// TIA Portal project "Industry 4.0_Plant_Logic" (V16) (continued)
REGION Network 1: Filling Process from Tank1
   // When bottle is detected at filling Station, after 2 sec, Tank 01 outlet valve is opened and Pump motor is started.
   // 
   // Tank 01 Outlet valve is closed when defined Liquid A percentage is filled in the bottle.
   // 
   // Liquid A filled value is then moved into Database for Storing purpose.
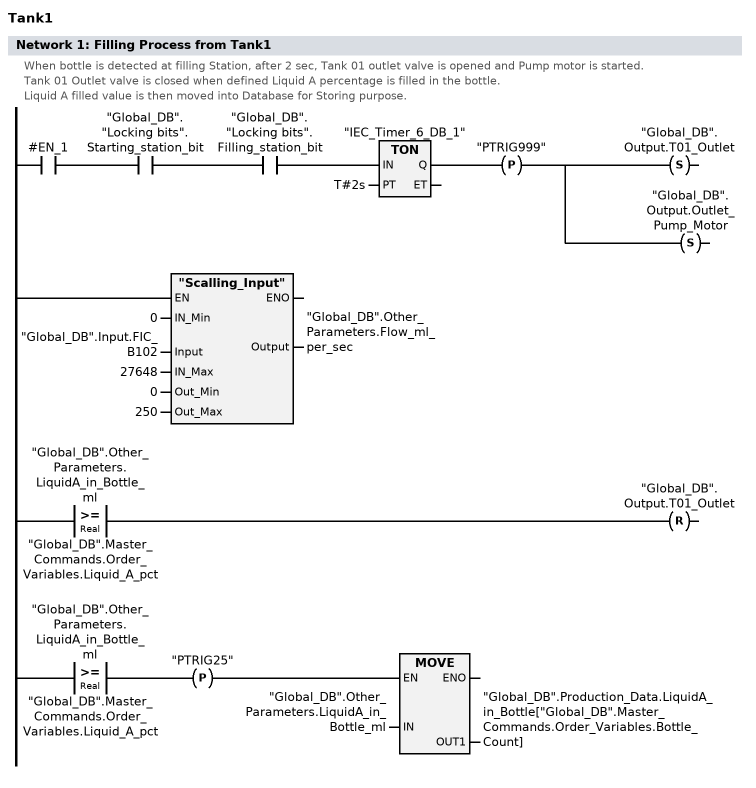
   "IEC_Timer_6_DB_1".TON(IN := #EN_1 AND "Global_DB"."Locking bits".Starting_station_bit AND "Global_DB"."Locking bits".Filling_station_bit,
                          PT := T#2s);
   #_w1 := "IEC_Timer_6_DB_1".Q AND NOT "PTRIG999";   // rising edge
   "PTRIG999" := "IEC_Timer_6_DB_1".Q;
   IF #_w1 THEN
       "Global_DB".Output.T01_Outlet := TRUE;
       "Global_DB".Output.Outlet_Pump_Motor := TRUE;
   END_IF;
   "Scalling_Input"(IN_Min := 0,
                    Input := "Global_DB".Input.FIC_B102,
                    IN_Max := 27648,
                    Out_Min := 0,
                    Out_Max := 250,
                    Output => "Global_DB".Other_Parameters.Flow_ml_per_sec);
   IF "Global_DB".Other_Parameters.LiquidA_in_Bottle_ml >= "Global_DB".Master_Commands.Order_Variables.Liquid_A_pct THEN
       "Global_DB".Output.T01_Outlet := FALSE;
   END_IF;
   #_w2 := "Global_DB".Other_Parameters.LiquidA_in_Bottle_ml >= "Global_DB".Master_Commands.Order_Variables.Liquid_A_pct;
   #_w3 := #_w2 AND NOT "PTRIG25";   // rising edge
   "PTRIG25" := #_w2;
   IF #_w3 THEN
       "Global_DB".Production_Data.LiquidA_in_Bottle["Global_DB".Master_Commands.Order_Variables.Bottle_Count] := "Global_DB".Other_Parameters.LiquidA_in_Bottle_ml;
   END_IF;
END_REGION
END_FUNCTION_BLOCK

FUNCTION_BLOCK "Tank2"   // FB5, LAD
{ S7_Optimized_Access := 'TRUE' }
VERSION : 0.1
   VAR_INPUT
      EN_2 : Bool;
   END_VAR
   VAR_TEMP   // added for the SCL form of the ladder/FBD networks
      _w1 : Bool;
      _w2 : Bool;
      _w3 : Bool;
   END_VAR
BEGIN

REGION Network 1: Tank02 Outlet Solenoid Valve
   // When bottle is filled with liquid A, after 3 sec, Tank 02 outlet valve is opened and Pump motor is started to fill liquid B.
   // 
   // Tank 02 Outlet valve is closed when defined Liquid B percentage is filled in the bottle.
   // 
   // Liquid B filled value is then moved into Database for Storing purpose.
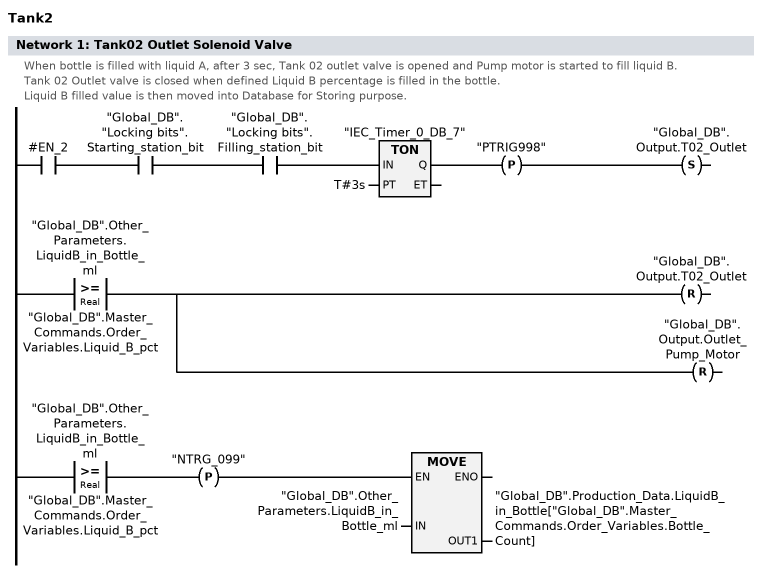
   "IEC_Timer_0_DB_7".TON(IN := #EN_2 AND "Global_DB"."Locking bits".Starting_station_bit AND "Global_DB"."Locking bits".Filling_station_bit,
                          PT := T#3s);
   #_w1 := "IEC_Timer_0_DB_7".Q AND NOT "PTRIG998";   // rising edge
   "PTRIG998" := "IEC_Timer_0_DB_7".Q;
   IF #_w1 THEN "Global_DB".Output.T02_Outlet := TRUE; END_IF;
   IF "Global_DB".Other_Parameters.LiquidB_in_Bottle_ml >= "Global_DB".Master_Commands.Order_Variables.Liquid_B_pct THEN
       "Global_DB".Output.T02_Outlet := FALSE;
       "Global_DB".Output.Outlet_Pump_Motor := FALSE;
   END_IF;
   #_w2 := "Global_DB".Other_Parameters.LiquidB_in_Bottle_ml >= "Global_DB".Master_Commands.Order_Variables.Liquid_B_pct;
   #_w3 := #_w2 AND NOT "NTRG_099";   // rising edge
   "NTRG_099" := #_w2;
   IF #_w3 THEN
       "Global_DB".Production_Data.LiquidB_in_Bottle["Global_DB".Master_Commands.Order_Variables.Bottle_Count] := "Global_DB".Other_Parameters.LiquidB_in_Bottle_ml;
   END_IF;
END_REGION
END_FUNCTION_BLOCK

FUNCTION_BLOCK "ProductionData_Reset"   // FB6, SCL
{ S7_Optimized_Access := 'TRUE' }
VERSION : 0.1
BEGIN

   // when number of filled bottles = Ordered bottle
   // reset the production data buffer and flag order completed To TRUE

   IF "Global_DB".Master_Commands.Order_Variables.Bottle_Count > "Global_DB".Master_Commands.Order_Variables.Quantity THEN
       FOR "Global_DB".Other_Parameters.index := 1 TO 5 BY 1 DO
           "Global_DB".Production_Data.Total_Liquid_in_Bottle["Global_DB".Other_Parameters.index] := 0.0;
           "Global_DB".Production_Data.LiquidA_in_Bottle["Global_DB".Other_Parameters.index] := 0.0;
           "Global_DB".Production_Data.LiquidB_in_Bottle["Global_DB".Other_Parameters.index] := 0.0;
       END_FOR;
       "Global_DB".Master_Commands.Order_Variables.Order_completed := True;
    END_IF;

    // when order is complete, reset the order data

   IF "Global_DB".Master_Commands.Order_Variables.Order_completed = True THEN
       "Global_DB".Master_Commands.Order_Variables.Bottle_Count := 1;
       "Global_DB".Master_Commands.Order_Variables.Order_ID := 0;
       "Global_DB".Master_Commands.Order_Variables.Quantity := 0;
       "Global_DB".Master_Commands.Order_Variables.Liquid_A_pct := 0;
       "Global_DB".Master_Commands.Order_Variables.Liquid_B_pct := 0;
       "Global_DB".Master_Commands.Order_Variables.Order_received := FALSE;
       // "Global_DB".Master_Commands.Order_Variables.Order_completed := FALSE;
   END_IF;
END_FUNCTION_BLOCK

FUNCTION_BLOCK "Reseting_order"   // FB7, SCL
{ S7_Optimized_Access := 'TRUE' }
VERSION : 0.1
BEGIN
   // when next order is received, turn Order_completed flag to FALSE

   "R_TRIG_DB"(CLK := "Global_DB".Master_Commands.Order_Variables.Order_received);

   IF "R_TRIG_DB".Q THEN
       "Global_DB".Master_Commands.Order_Variables.Order_completed := FALSE;
   END_IF;
END_FUNCTION_BLOCK

FUNCTION_BLOCK "Operation_cycle"   // FB8, LAD
{ S7_Optimized_Access := 'TRUE' }
VERSION : 0.1
   VAR
      begun : Bool;
   END_VAR
   VAR_TEMP
      ons1 : Bool;
   END_VAR
   VAR_TEMP   // added for the SCL form of the ladder/FBD networks
      _w1 : Bool;
      _w2 : Bool;
      _w3 : Bool;
   END_VAR
BEGIN

REGION Network 1: Calculate Operation time for one bottle filling and storing in Database for every bottle
   // Operation begin - robot has picked bottle
   // Operation finished - bottle if capped and placed by robot
   // 
   // Note : currently these variables are not getting real-feedback from robots. These are for just simulation.
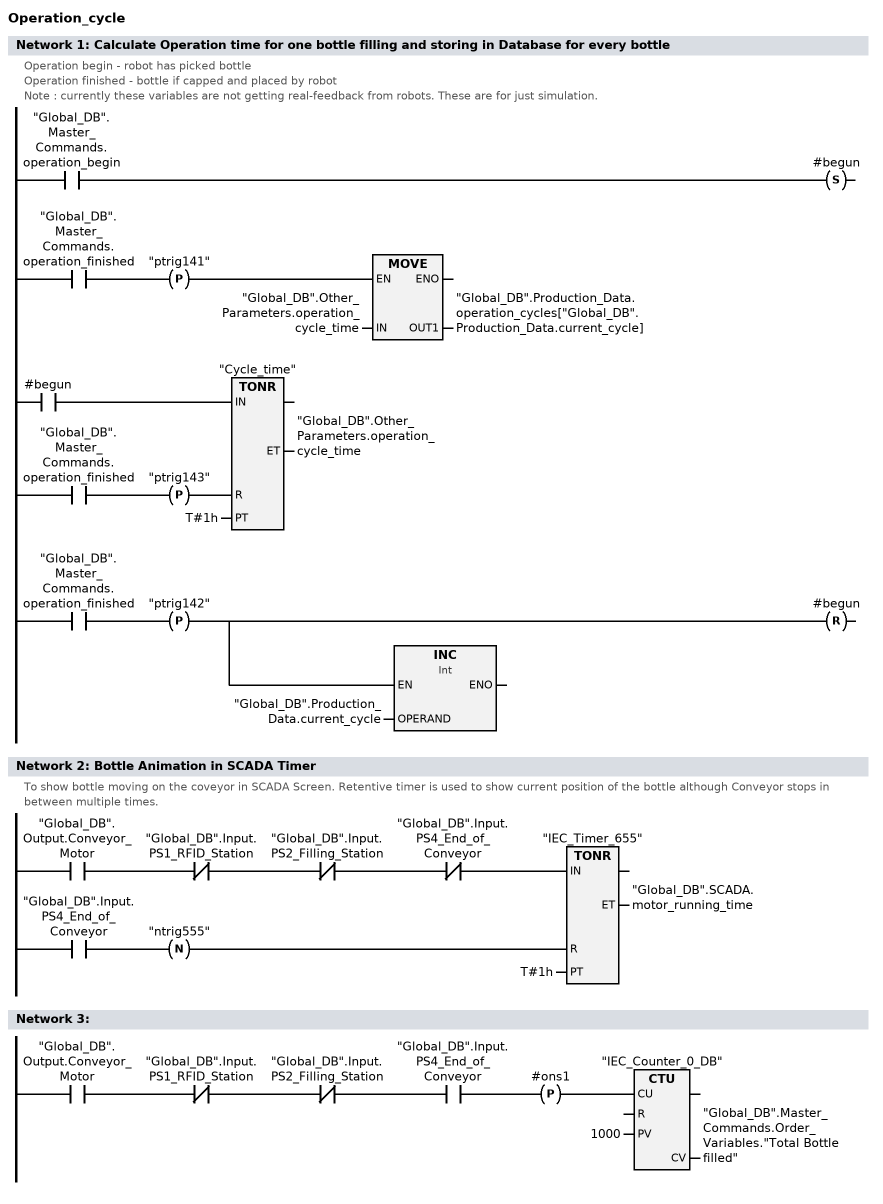
   IF "Global_DB".Master_Commands.operation_begin THEN #begun := TRUE; END_IF;
   #_w1 := "Global_DB".Master_Commands.operation_finished AND NOT "ptrig141";   // rising edge
   "ptrig141" := "Global_DB".Master_Commands.operation_finished;
   IF #_w1 THEN
       "Global_DB".Production_Data.operation_cycles["Global_DB".Production_Data.current_cycle] := "Global_DB".Other_Parameters.operation_cycle_time;
   END_IF;
   #_w2 := "Global_DB".Master_Commands.operation_finished AND NOT "ptrig143";   // rising edge
   "ptrig143" := "Global_DB".Master_Commands.operation_finished;
   "Cycle_time".TONR(IN := #begun,
                     R := #_w2,
                     PT := T#1h,
                     ET => "Global_DB".Other_Parameters.operation_cycle_time);
   #_w3 := "Global_DB".Master_Commands.operation_finished AND NOT "ptrig142";   // rising edge
   "ptrig142" := "Global_DB".Master_Commands.operation_finished;
   IF #_w3 THEN
       #begun := FALSE;
       "Global_DB".Production_Data.current_cycle := "Global_DB".Production_Data.current_cycle + 1;
   END_IF;
END_REGION

REGION Network 2: Bottle Animation in SCADA Timer
   // To show bottle moving on the coveyor in SCADA Screen. Retentive timer is used to show current position of the bottle although Conveyor stops in between multiple times.
   #_w1 := NOT "Global_DB".Input.PS4_End_of_Conveyor AND "ntrig555";   // falling edge
   "ntrig555" := "Global_DB".Input.PS4_End_of_Conveyor;
   "IEC_Timer_655".TONR(IN := "Global_DB".Output.Conveyor_Motor AND NOT "Global_DB".Input.PS1_RFID_Station AND NOT "Global_DB".Input.PS2_Filling_Station AND NOT "Global_DB".Input.PS4_End_of_Conveyor,
                        R := #_w1,
                        PT := T#1h,
                        ET => "Global_DB".SCADA.motor_running_time);
END_REGION

REGION Network 3
   #_w1 := "Global_DB".Output.Conveyor_Motor AND NOT "Global_DB".Input.PS1_RFID_Station AND NOT "Global_DB".Input.PS2_Filling_Station AND "Global_DB".Input.PS4_End_of_Conveyor;
   #_w2 := #_w1 AND NOT #ons1;   // rising edge
   #ons1 := #_w1;
   "IEC_Counter_0_DB".CTU(CU := #_w2,
                          PV := 1000,
                          CV => "Global_DB".Master_Commands.Order_Variables."Total Bottle filled");
END_REGION
END_FUNCTION_BLOCK

FUNCTION_BLOCK "Array_Voltage_Logic"   // FB9, SCL
{ S7_Optimized_Access := 'TRUE' }
VERSION : 0.1
BEGIN




       "Global_DB".Array_Voltage["i"] :="Global_DB".Motor_Output_PCT;
       "i" := "i" + 1;
END_FUNCTION_BLOCK

// folder: Functions

FUNCTION "Scalling_Input" : Void   // FC1, FBD
{ S7_Optimized_Access := 'TRUE' }
VERSION : 0.1
   VAR_INPUT
      IN_Min : Int;
      Input : Int;
      IN_Max : Int;
      Out_Min : Int;
      Out_Max : Int;
   END_VAR
   VAR_OUTPUT
      Output : Real;
   END_VAR
   VAR_TEMP
      Normed : Real;
   END_VAR
BEGIN

REGION Network 1
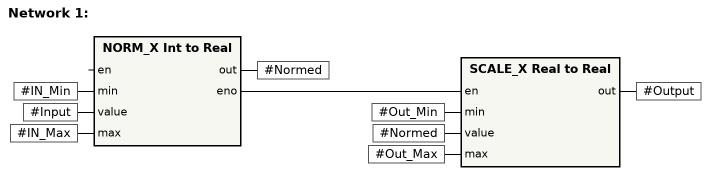
   #Normed := NORM_X(MIN := #IN_Min, VALUE := #Input, MAX := #IN_Max);
   #Output := SCALE_X(MIN := #Out_Min, VALUE := #Normed, MAX := #Out_Max);
END_REGION
END_FUNCTION

FUNCTION "Scalling_Output" : Void   // FC2, FBD
{ S7_Optimized_Access := 'TRUE' }
VERSION : 0.1
   VAR_INPUT
      IN_Min : Int;
      Input : Int;
      IN_Max : Int;
      Out_Min : Int;
      Out_Max : Int;
   END_VAR
   VAR_OUTPUT
      Output : Int;
   END_VAR
   VAR_TEMP
      Normed : Real;
   END_VAR
BEGIN

REGION Network 1
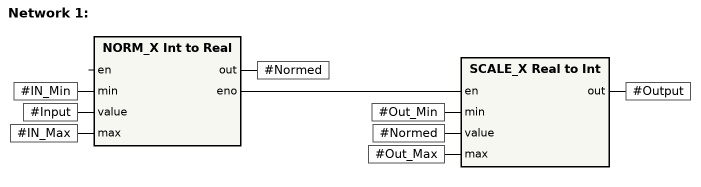
   #Normed := NORM_X(MIN := #IN_Min, VALUE := #Input, MAX := #IN_Max);
   #Output := SCALE_X(MIN := #Out_Min, VALUE := #Normed, MAX := #Out_Max);
END_REGION
END_FUNCTION

FUNCTION "Reading" : Void   // FC3, SCL
{ S7_Optimized_Access := 'TRUE' }
VERSION : 0.1
BEGIN
   // Reading inputs from PLC terminals to Global_DB

   "Global_DB".Input.FIC_B102 := "FIC_B102";
   "Global_DB".Input.LIC_B101 := "LIC_B101";
   "Global_DB".Input.PS1_RFID_Station := "PS1_RFID_Station";
   "Global_DB".Input.PS2_Filling_Station := "PS2_Filling_Station";
   "Global_DB".Input.PS3_Quality_Station := "PS3_Quality_Station";
   "Global_DB".Input.PS4_End_of_Conveyor := "PS4_End_of_Conveyor";
   "Global_DB".Input.T01_Low_Level := "T01_Low_Level";
   "Global_DB".Input.T01_High_Level := "T01_High_Level";
END_FUNCTION

FUNCTION "Writing" : Void   // FC4, SCL
{ S7_Optimized_Access := 'TRUE' }
VERSION : 0.1
BEGIN
   // Writing Output from Global_DB to PLC Terminal

   "T01_Outlet" := "Global_DB".Output.T01_Outlet;
   "T02_Outlet" := "Global_DB".Output.T02_Outlet;

   "Outlet_Pump_Motor" := "Global_DB".Output.Outlet_Pump_Motor;
   "Conveyor_Motor" := "Global_DB".Output.Conveyor_Motor;
END_FUNCTION

FUNCTION "Filling_Logik" : Void   // FC5, LAD
{ S7_Optimized_Access := 'TRUE' }
VERSION : 0.1
   VAR_INPUT
      PS2_Filling_Station : Bool;
      FIC_B102 : Int;
      Liquid_AorB_in_Bottle_ml : Real;
      Liquid_AorB_pct : Int;
      Wait_to_fill : Time;
   END_VAR
   VAR_OUTPUT
      Flow_ml_per_sec : Real;
      FillingData_LiqAorB_ml : Real;
   END_VAR
   VAR_IN_OUT
      Outlet_of_tanks : Bool;
   END_VAR
   VAR_TEMP
      PTRIG1 : Bool;
      PTRIG2 : Bool;
      PTRIG3 : Bool;
      PTRIG4 : Bool;
   END_VAR
BEGIN

REGION Network 1
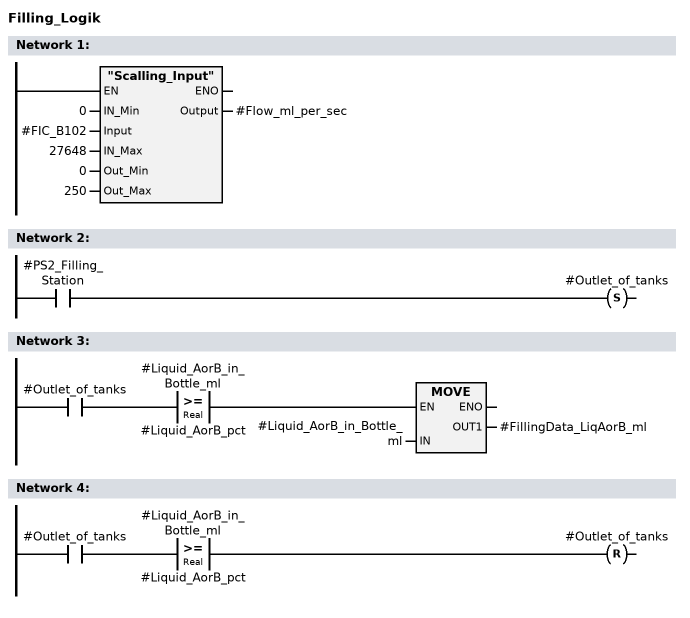
   RUNG wire#powerrail
      "Scalling_Input"(IN_Min := 0, Input := #FIC_B102, IN_Max := 27648, Out_Min := 0, Out_Max := 250, Output => #Flow_ml_per_sec)
   END_RUNG
   // the same network as SCL:
   "Scalling_Input"(IN_Min := 0,
                    Input := #FIC_B102,
                    IN_Max := 27648,
                    Out_Min := 0,
                    Out_Max := 250,
                    Output => #Flow_ml_per_sec);
END_REGION

REGION Network 2
   RUNG wire#powerrail
      Contact( #PS2_Filling_Station )
      S_Coil( #Outlet_of_tanks )
   END_RUNG
   // the same network as SCL:
   IF #PS2_Filling_Station THEN #Outlet_of_tanks := TRUE; END_IF;
END_REGION

REGION Network 3
   RUNG wire#powerrail
      Contact( #Outlet_of_tanks )
      { S7_Templates := "SrcType := Real" } GE_Contact(in1 := #Liquid_AorB_in_Bottle_ml, in2 := #Liquid_AorB_pct)
      Move(in := #Liquid_AorB_in_Bottle_ml, out1 => #FillingData_LiqAorB_ml)
   END_RUNG
   // the same network as SCL:
   IF #Outlet_of_tanks AND (#Liquid_AorB_in_Bottle_ml >= #Liquid_AorB_pct) THEN
       #FillingData_LiqAorB_ml := #Liquid_AorB_in_Bottle_ml;
   END_IF;
END_REGION

REGION Network 4
   RUNG wire#powerrail
      Contact( #Outlet_of_tanks )
      { S7_Templates := "SrcType := Real" } GE_Contact(in1 := #Liquid_AorB_in_Bottle_ml, in2 := #Liquid_AorB_pct)
      R_Coil( #Outlet_of_tanks )
   END_RUNG
   // the same network as SCL:
   IF #Outlet_of_tanks AND (#Liquid_AorB_in_Bottle_ml >= #Liquid_AorB_pct) THEN
       #Outlet_of_tanks := FALSE;
   END_IF;
END_REGION
END_FUNCTION

(* ===== HMI "HMI_RT_1" =====
system functions are stored by id; their names below are inferred from use
connection "PLCs71200": ETHERNET, SMART_S7_1200_OMS
connection "HMI_Connection_1": ETHERNET, SMART_S7_1200_OMS

HMI tags "Default tag table"
   "Conveyor_Motor" : Bool = PLC Global_DB.Output.Conveyor_Motor AT %DB1.DBX6.3, 1 s
   "Outlet_Pump_Motor" : Bool = PLC Global_DB.Output.Outlet_Pump_Motor AT %DB1.DBX6.2, 1 s
   "T01_Outlet_Valve" : Bool = PLC Global_DB.Output.T01_Outlet AT %DB1.DBX6.0, 1 s
   "T02_Outlet_Valve" : Bool = PLC Global_DB.Output.T02_Outlet AT %DB1.DBX6.1, 1 s
   "T02_fluid Low level" : Real = PLC Global_DB.Other_Parameters.T02_Low_Level_Limit AT %DB1.DBD30, 1 s
   "Global_DB_Other_Parameters_Liquid_A_pct" : Int = PLC Global_DB.Master_Commands.Order_Variables.Liquid_A_pct AT %DB1.DBW52, 1 s
   "Global_DB_Other_Parameters_Liquid_B_pct" : Int = PLC Global_DB.Master_Commands.Order_Variables.Liquid_B_pct AT %DB1.DBW54, 1 s
   "Total_Liquid_in_Bottle{0}" : Array [0..4] of Real = PLC Global_DB.Production_Data.Total_Liquid_in_Bottle AT %DB1.DBX66.0, 1 s
   "T02_Low_Level_Limit" : Real = PLC Global_DB.Other_Parameters.T02_Low_Level_Limit AT %DB1.DBD30, 1 s
   "Global_DB_Input_T01_Low_Level" : Bool = PLC Global_DB.Input.T01_Low_Level AT %DB1.DBX4.4, 1 s
   "Global_DB_Input_T01_High_Level" : Bool = PLC Global_DB.Input.T01_High_Level AT %DB1.DBX4.5, 1 s
   "Error_Alarm" : Word = PLC Global_DB.Error.Alarm AT %DB1.DBW42, 1 s
   "Global_DB_Input_FIC_B102" : Int = PLC Global_DB.Input.FIC_B102 AT %DB1.DBW0, 1 s
   "Global_DB_Input_LIC_B101" : Int = PLC Global_DB.Input.LIC_B101 AT %DB1.DBW2, 1 s
   "Global_DB_Production_Data_Bottle_Count" : Int = PLC Global_DB.Master_Commands.Order_Variables.Bottle_Count AT %DB1.DBW58, 1 s
   "Flow_ml_per_sec" : Real = PLC Global_DB.Other_Parameters.Flow_ml_per_sec AT %DB1.DBD10, 1 s
   "PS1_RFID_Station" : Bool = PLC Global_DB.Input.PS1_RFID_Station AT %DB1.DBX4.0, 1 s
   "PS2_Filling_Station" : Bool = PLC Global_DB.Input.PS2_Filling_Station AT %DB1.DBX4.1, 1 s
   "PS3_Quality_Station" : Bool = PLC Global_DB.Input.PS3_Quality_Station AT %DB1.DBX4.2, 1 s
   "PS4_End_of_Conveyor" : Bool = PLC Global_DB.Input.PS4_End_of_Conveyor AT %DB1.DBX4.3, 1 s

discrete alarms
   1: 'Level of Tank01 is high', class Errors, trigger "Global_DB_Error_HIgh level Alarm T01" bit 0
   2: 'Level of Tank01 is low', class Errors, trigger "Global_DB_Error_low level Alarm T01" bit 0

analog alarms
   4: 'Level of Tank02 is high', class Warnings, trigger "Global_DB_Other_Parameters_T02_High_Level_Limit"
   5: 'Level of Tank02 is low', class Warnings, trigger "T02_Low_Level_Limit"

recipe "combinations": Liquid A <- "Global_DB_Other_Parameters_Liquid_A_pct", Liquid B <- "Global_DB_Other_Parameters_Liquid_B_pct"

screen "Different jobs" 800x480
   TextField "Text field_1" at 339,11 size 221x27; Text 'Diffrent Jobs / Gruppe der Ingenieure'
   GraphicView "Graphic view_61" at 2,4 size 149x43; Picture "logo2"
   DateTimeField "Date/time field_1" at 629,14 size 166x19
   Button "Back" at 181,104 size 188x64; TextOn 'Back / Zurück'; TextOff 'Back / Zurück'
      on Release: function_efd93a16()
   Button "Toggle language" at 177,208 size 192x70; TextOn 'Toggle language / Sprache Wechseln'; TextOff 'Toggle language / Sprache Wechseln'
      on Release: function_fb9197e8(-1)
   Button "Online" at 177,320 size 192x66; TextOn 'Online'; TextOff 'Online'
   Button "Offline" at 460,103 size 189x65; TextOn 'Offline'; TextOff 'Offline'
   Button "Stop Runtime" at 460,209 size 189x69; TextOn 'Stop Runtime / Laufzeit anhalten'; TextOff 'Stop Runtime / Laufzeit anhalten'
   Button "Transfer" at 457,320 size 192x65; TextOn 'Transfer / Übertragung'; TextOff 'Transfer / Übertragung'
   Button "Button_1" at 6,432 size 88x38; TextOff 'Root'
      on Release: ActivateScreen("Root screen", 0)
      on Press: ActivateScreen("Root screen", 0)
   Button "Button_2" at 99,432 size 93x38; TextOff 'User / Benutzer'
      on Release: ActivateScreen("User administration", 0)
      on Press: ActivateScreen("User administration", 0)
   Button "Button_3" at 197,431 size 96x39; TextOff 'Alarms / Alarme'
      on Release: ActivateScreen("Alarm screen", 0)
      on Press: ActivateScreen("Alarm screen", 0)
   Button "Button_4" at 298,431 size 121x39; TextOff 'PLC diagnose / SPS Diagnose'
      on Release: ActivateScreen("SIMATIC PLC system diagnostics", 0)
      on Press: ActivateScreen("SIMATIC PLC system diagnostics", 0)
   Button "Button_5" at 425,431 size 106x39; TextOff 'Recipes / Rezepte'
      on Release: ActivateScreen("Recipes management", 0)
      on Press: ActivateScreen("Recipes management", 0)
   Button "Button_6" at 537,431 size 113x39; TextOff 'Visulization / Visulisierung'
      on Release: ActivateScreen("visualization", 0)
      on Press: ActivateScreen("visualization", 0)
   Button "Button_7" at 654,431 size 139x39; TextOff 'Historic Data / Frühere Daten'
      on Release: ActivateScreen("Historical Data", 0)
      on Press: ActivateScreen("Historical Data", 0)

screen "visualization" 800x480
   GraphicView "Graphic view_38" at 637,99 size 155x90; Picture "Graphic_80"
   GraphicView "Graphic view_91" at 719,110 size 19x17; Picture "Graphic_70"
   GraphicView "Graphic view_84" at 735,110 size 19x17; Picture "Graphic_70"
   GraphicView "Graphic view_26" at 751,110 size 19x17; Picture "Graphic_70"
   GraphicView "Graphic view_83" at 768,110 size 19x17; Picture "Graphic_70"
   TextField "Text field_2" at 600,134 size 15x23; Text '4'
   GraphicView "Graphic view_22" at 285,216 size 38x24; Picture "Graphic_43"
   GraphicView "Graphic view_4" at 442,213 size 29x22; Picture "Graphic_60"
   GraphicView "Graphic view_32" at 2,111 size 162x71; Picture "Graphic_76"
   GraphicView "Graphic view_27" at 181,310 size 49x14; Picture "Graphic_65"
   GraphicView "Graphic view_61" at 2,4 size 149x43; Picture "logo2"
   DateTimeField "Date/time field_1" at 629,14 size 167x19
   TextField "Text field_1" at 346,11 size 115x25; Text 'Visulization / Visulisierung'
   Group "Group_1" at 637,99 size 155x90; Picture "Graphic_80"
   GraphicView "Graphic view_72" at 633,201 size 162x71; Picture "Graphic_76"
   GraphicView "Graphic view_82" at 713,205 size 22x17; Picture "Graphic_70"
   GraphicView "Graphic view_85" at 676,205 size 22x17; Picture "Graphic_70"
   GraphicView "Graphic view_87" at 694,205 size 22x17; Picture "Graphic_70"
   GraphicView "Graphic view_93" at 690,211 size 22x17; Picture "Graphic_70"
   GraphicView "Graphic view_103" at 671,211 size 22x17; Picture "Graphic_70"
   Group "Group_4" at 587,131 size 43x28
   GraphicView "Graphic view_89" at 658,205 size 22x17; Picture "Graphic_70"
   GraphicView "Graphic view_86" at 653,211 size 22x17; Picture "Graphic_70"
   GraphicView "Graphic view_92" at 649,217 size 22x17; Picture "Graphic_70"
   GraphicView "Graphic view_90" at 645,222 size 22x17; Picture "Graphic_70"
   GraphicView "Graphic view_80" at 708,211 size 22x17; Picture "Graphic_70"
   GraphicView "Graphic view_1" at 258,95 size 95x94; Picture "Graphic_1"
   GraphicView "Graphic view_21" at 318,221 size 130x14; Picture "Graphic_41"
   GraphicView "Graphic view_2" at 414,97 size 95x94; Picture "Graphic_1"
   GraphicView "Graphic view_11" at 415,100 size 28x90; Picture "Graphic_15"
   GraphicView "Graphic view_12" at 451,187 size 22x16; Picture "Graphic_57"
   GraphicView "Graphic view_19" at 451,201 size 32x16; Picture "Graphic_48"
      Appearance <- "T01_Outlet_Valve"
   GraphicView "Graphic view_5" at 280,61 size 41x122; Picture "Graphic_4"
   GraphicView "Graphic view_9" at 322,236 size 44x38; Picture "Graphic_9"
   GraphicView "Graphic view_7" at 240,214 size 54x28; Picture "Graphic_10"
      Appearance <- "Outlet_Pump_Motor"
   GraphicView "Graphic view_13" at 292,185 size 24x17; Picture "Graphic_57"
   GraphicView "Graphic view_18" at 292,200 size 35x19; Picture "Graphic_48"
      Appearance <- "T02_Outlet_Valve"
   GraphicView "Graphic view_23" at 294,237 size 20x12; Picture "Graphic_57"
   GraphicView "Graphic view_24" at 364,257 size 18x17; Picture "Graphic_63"
   GraphicView "Graphic view_28" at 391,282 size 22x22; Picture "Graphic_72"
   GraphicView "Graphic view_25" at 377,257 size 36x27; Picture "Graphic_64"
   GraphicView "Graphic view_20" at 294,247 size 32x27; Picture "Graphic_62"
   GraphicView "Graphic view_6" at 486,102 size 47x25; Picture "Graphic_5"
      Appearance <- "Global_DB_Input_T01_High_Level"
   GraphicView "Graphic view_8" at 486,170 size 47x25; Picture "Graphic_5"
      Appearance <- "Global_DB_Input_T01_Low_Level"
   IOField "I/O field_1" at 563,220 size 71x32; FormatPattern 999
      ProcessValue <- "Global_DB_Production_Data_Bottle_Count"
   IOField "I/O field_2" at 102,246 size 102x32; FormatPattern 999.99; Unit ml/s
      ProcessValue <- "Flow_ml_per_sec"
   GraphicView "Graphic view_33" at 100,114 size 22x17; Picture "Graphic_70"
   GraphicView "Graphic view_34" at 95,121 size 22x17; Picture "Graphic_70"
   GraphicView "Graphic view_35" at 82,114 size 22x17; Picture "Graphic_70"
   GraphicView "Graphic view_36" at 45,113 size 22x17; Picture "Graphic_70"
   GraphicView "Graphic view_37" at 28,113 size 22x17; Picture "Graphic_70"
   GraphicView "Graphic view_39" at 65,113 size 22x17; Picture "Graphic_70"
   GraphicView "Graphic view_41" at 22,119 size 22x17; Picture "Graphic_70"
   GraphicView "Graphic view_42" at 76,121 size 22x17; Picture "Graphic_70"
   GraphicView "Graphic view_43" at 41,118 size 22x17; Picture "Graphic_70"
   GraphicView "Graphic view_44" at 60,119 size 22x17; Picture "Graphic_70"
   GraphicView "Graphic view_46" at 118,115 size 22x17; Picture "Graphic_70"
   GraphicView "Graphic view_47" at 72,127 size 22x17; Picture "Graphic_70"
   GraphicView "Graphic view_51" at 53,127 size 22x17; Picture "Graphic_70"
   TextField "Text field_4" at 176,132 size 25x23; Text '6 / 14'
   GraphicView "Graphic view_50" at 36,126 size 22x17; Picture "Graphic_70"
   GraphicView "Graphic view_48" at 30,132 size 22x17; Picture "Graphic_70"
   GraphicView "Graphic view_49" at 17,126 size 22x17; Picture "Graphic_70"
   GraphicView "Graphic view_45" at 13,132 size 22x17; Picture "Graphic_70"
   TextField "Text field_3" at 8,250 size 93x23; Text 'Flow Rate:'
   GraphicView "Graphic view_10" at 260,98 size 28x90; Picture "Graphic_15"
   Button "Button_1" at 6,432 size 88x38; TextOff 'Root'
      on Release: ActivateScreen("Root screen", 0)
      on Press: ActivateScreen("Root screen", 0)
   Button "Button_2" at 99,432 size 93x38; TextOff 'User / Benutzer'
      on Release: ActivateScreen("User administration", 0)
      on Press: ActivateScreen("User administration", 0)
   Button "Button_3" at 197,431 size 96x39; TextOff 'Alarms / Alarme'
      on Release: ActivateScreen("Alarm screen", 0)
      on Press: ActivateScreen("Alarm screen", 0)
   Button "Button_4" at 298,431 size 121x39; TextOff 'PLC diagnose / SPS Diagnose'
      on Release: ActivateScreen("SIMATIC PLC system diagnostics", 0)
      on Press: ActivateScreen("SIMATIC PLC system diagnostics", 0)
   Button "Button_5" at 425,431 size 106x39; TextOff 'Recipes / Rezepte'
      on Release: ActivateScreen("Recipes management", 0)
      on Press: ActivateScreen("Recipes management", 0)
   Button "Button_6" at 537,431 size 113x39; TextOff 'Visulization / Visulisierung'
      on Release: ActivateScreen("visualization", 0)
      on Press: ActivateScreen("visualization", 0)
   Button "Button_7" at 654,431 size 139x39; TextOff 'Historic Data / Frühere Daten'
      on Release: ActivateScreen("Historical Data", 0)
      on Press: ActivateScreen("Historical Data", 0)
   GraphicView "Graphic view_68" at 140,388 size 41x27; Picture "Graphic_93"
      Appearance <- "Conveyor_Motor"
   GraphicView "Graphic view_17" at 137,331 size 510x69; Picture "Graphic_28"
   GraphicView "Graphic view_40" at 185,338 size 35x24; Picture "Graphic_88"
   GraphicView "Graphic view_29" at 241,304 size 29x72; Picture "Graphic_70"
      Visibility <- "PS1_RFID_Station"
   GraphicView "Graphic view_15" at 265,306 size 22x41; Picture "Graphic_24"
      Appearance <- "PS1_RFID_Station"
   GraphicView "Graphic view_67" at 323,304 size 29x72; Picture "Graphic_70"
      Visibility <- "PS2_Filling_Station"
   GraphicView "Graphic view_14" at 340,305 size 22x41; Picture "Graphic_24"
      Appearance <- "PS2_Filling_Station"
   GraphicView "Graphic view_3" at 445,307 size 22x41; Picture "Graphic_24"
      Appearance <- "PS3_Quality_Station"
   GraphicView "Graphic view_65" at 423,304 size 29x72; Picture "Graphic_70"
      Visibility <- "PS3_Quality_Station"
   GraphicView "Graphic view_63" at 511,304 size 29x72; Picture "Graphic_70"
      Visibility <- "PS4_End_of_Conveyor"
   GraphicView "Graphic view_16" at 532,307 size 22x41; Picture "Graphic_24"
      Appearance <- "PS4_End_of_Conveyor"

screen "Root screen" 800x480
   TextField "HmiScreenItemData" at 64,85 size 675x54; Text 'Welcome to liquid filling plant based on Industry 4.0 / Willkommen bei der Flüssigkeitsabfüllanlage auf Basis von Industrie 4.0'
   TextField "Text field_1" at 339,10 size 158x27; Text 'Root Screen / Root Bildschirm'
   GraphicView "Graphic view_61" at 2,4 size 149x43; Picture "logo2"
   DateTimeField "Date/time field_1" at 629,14 size 166x19
   Button "Button_8" at 263,167 size 115x69; TextOff 'START'
   Button "Button_9" at 425,166 size 115x69; TextOff 'STOP / STOPP'
   Switch "Switch_1" at 287,262 size 226x63; TextOn 'Emergency is pressed / Notruf wird gedrückt'; CaptionText 'Switch'; TextOff 'Emergency is released / Notfall wird ausgelöst'
   Button "Button_1" at 6,432 size 88x38; TextOff 'Root'
      on Release: ActivateScreen("Root screen", 0)
      on Press: ActivateScreen("Root screen", 0)
   Button "Button_2" at 99,432 size 93x38; TextOff 'User / Benutzer'
      on Release: ActivateScreen("User administration", 0)
      on Press: ActivateScreen("User administration", 0)
   Button "Button_3" at 197,431 size 96x39; TextOff 'Alarms / Alarme'
      on Release: ActivateScreen("Alarm screen", 0)
      on Press: ActivateScreen("Alarm screen", 0)
   Button "Button_4" at 298,431 size 121x39; TextOff 'PLC diagnose / SPS Diagnose'
      on Release: ActivateScreen("SIMATIC PLC system diagnostics", 0)
      on Press: ActivateScreen("SIMATIC PLC system diagnostics", 0)
   Button "Button_5" at 425,431 size 106x39; TextOff 'Recipes / Rezepte'
      on Release: ActivateScreen("Recipes management", 0)
      on Press: ActivateScreen("Recipes management", 0)
   Button "Button_6" at 537,431 size 113x39; TextOff 'Visulization / Visulisierung'
      on Release: ActivateScreen("visualization", 0)
      on Press: ActivateScreen("visualization", 0)
   Button "Button_7" at 654,431 size 139x39; TextOff 'Historic Data / Frühere Daten'
      on Release: ActivateScreen("Historical Data", 0)
      on Press: ActivateScreen("Historical Data", 0)
   Button "Button_12" at 9,156 size 176x46; TextOff 'Different Jobs / System Bildschirme'
      on Release: ActivateScreen("Different jobs", 0)
      on Press: ActivateScreen("Different jobs", 0)
   Button "Button_11" at 16,222 size 157x45; TextOff 'Engineer / Ingenieur'; Authorization "Engineer"
      on Release: ActivateScreen("Engineer Screen", 0)
      on Press: ActivateScreen("Engineer Screen", 0)
   Button "Button_13" at 12,287 size 164x49; TextOff 'Change Langauge / Sprache Wechseln'
      on Click: function_fb9197e8(-1)

screen "User administration" 800x480
   TextField "Text field_1" at 319,10 size 198x27; Text 'User Administration / Benutzerverwaltung'
   GraphicView "Graphic view_61" at 2,4 size 149x43; Picture "logo2"
   DateTimeField "Date/time field_1" at 628,14 size 167x19
   UserView "User view_1" at 9,64 size 781x289
   Button "Button_8" at 10,372 size 134x39; TextOff 'Logoff / Abmeldung'
      on Release: function_f23ef4c9()
      on Press: function_f23ef4c9()
   Button "Button_1" at 6,432 size 88x38; TextOff 'Root'
      on Release: ActivateScreen("Root screen", 0)
      on Press: ActivateScreen("Root screen", 0)
   Button "Button_2" at 99,432 size 93x38; TextOff 'User / Benutzer'
      on Release: ActivateScreen("User administration", 0)
      on Press: ActivateScreen("User administration", 0)
   Button "Button_3" at 197,431 size 96x39; TextOff 'Alarms / Alarme'
      on Release: ActivateScreen("Alarm screen", 0)
      on Press: ActivateScreen("Alarm screen", 0)
   Button "Button_4" at 298,431 size 121x39; TextOff 'PLC diagnose / SPS Diagnose'
      on Release: ActivateScreen("SIMATIC PLC system diagnostics", 0)
      on Press: ActivateScreen("SIMATIC PLC system diagnostics", 0)
   Button "Button_5" at 425,431 size 106x39; TextOff 'Recipes / Rezepte'
      on Release: ActivateScreen("Recipes management", 0)
      on Press: ActivateScreen("Recipes management", 0)
   Button "Button_6" at 537,431 size 113x39; TextOff 'Visulization / Visulisierung'
      on Release: ActivateScreen("visualization", 0)
      on Press: ActivateScreen("visualization", 0)
   Button "Button_7" at 654,431 size 139x39; TextOff 'Historic Data / Frühere Daten'
      on Release: ActivateScreen("Historical Data", 0)
      on Press: ActivateScreen("Historical Data", 0)

screen "SIMATIC PLC system diagnostics" 800x480
   SysDiagControl "HmiScreenItemData" at 19,64 size 759x349
   TextField "Text field_1" at 314,9 size 224x27; Text 'PLC System Diagnostic / SPS Diagnose'
   GraphicView "Graphic view_61" at 2,4 size 149x43; Picture "logo2"
   DateTimeField "Date/time field_1" at 628,14 size 167x19
   Button "Button_1" at 6,432 size 88x38; TextOff 'Root'
      on Release: ActivateScreen("Root screen", 0)
      on Press: ActivateScreen("Root screen", 0)
   Button "Button_2" at 99,432 size 93x38; TextOff 'User / Benutzer'
      on Release: ActivateScreen("User administration", 0)
      on Press: ActivateScreen("User administration", 0)
   Button "Button_3" at 197,431 size 96x39; TextOff 'Alarms / Alarme'
      on Release: ActivateScreen("Alarm screen", 0)
      on Press: ActivateScreen("Alarm screen", 0)
   Button "Button_4" at 298,431 size 121x39; TextOff 'PLC diagnose / SPS Diagnose'
      on Release: ActivateScreen("SIMATIC PLC system diagnostics", 0)
      on Press: ActivateScreen("SIMATIC PLC system diagnostics", 0)
   Button "Button_5" at 425,431 size 106x39; TextOff 'Recipes / Rezepte'
      on Release: ActivateScreen("Recipes management", 0)
      on Press: ActivateScreen("Recipes management", 0)
   Button "Button_6" at 537,431 size 113x39; TextOff 'Visulization / Visulisierung'
      on Release: ActivateScreen("visualization", 0)
      on Press: ActivateScreen("visualization", 0)
   Button "Button_7" at 654,431 size 139x39; TextOff 'Historic Data / Frühere Daten'
      on Release: ActivateScreen("Historical Data", 0)
      on Press: ActivateScreen("Historical Data", 0)

screen "Historical Data" 800x480
   on ClearScreen: function_efd5fb8c()
   TextField "Text field_1" at 339,10 size 175x27; Text 'Historical Data / Historische Daten'
   GraphicView "Graphic view_61" at 2,4 size 149x43; Picture "logo2"
   DateTimeField "Date/time field_1" at 628,14 size 167x19
   TrendView "Trend view_1" at 27,51 size 754x374
   Button "Button_1" at 6,432 size 88x38; TextOff 'Root'
      on Release: ActivateScreen("Root screen", 0)
      on Press: ActivateScreen("Root screen", 0)
   Button "Button_2" at 99,432 size 93x38; TextOff 'User / Benutzer'
      on Release: ActivateScreen("User administration", 0)
      on Press: ActivateScreen("User administration", 0)
   Button "Button_3" at 197,431 size 96x39; TextOff 'Alarms / Alarme'
      on Release: ActivateScreen("Alarm screen", 0)
      on Press: ActivateScreen("Alarm screen", 0)
   Button "Button_4" at 298,431 size 121x39; TextOff 'PLC diagnose / SPS Diagnose'
      on Release: ActivateScreen("SIMATIC PLC system diagnostics", 0)
      on Press: ActivateScreen("SIMATIC PLC system diagnostics", 0)
   Button "Button_5" at 425,431 size 106x39; TextOff 'Recipes / Rezepte'
      on Release: ActivateScreen("Recipes management", 0)
      on Press: ActivateScreen("Recipes management", 0)
   Button "Button_6" at 537,431 size 113x39; TextOff 'Visulization / Visulisierung'
      on Release: ActivateScreen("visualization", 0)
      on Press: ActivateScreen("visualization", 0)
   Button "Button_7" at 654,431 size 139x39; TextOff 'Historic Data / Frühere Daten'
      on Release: ActivateScreen("Historical Data", 0)
      on Press: ActivateScreen("Historical Data", 0)

screen "Recipes management" 800x480
   RecipeView "Recipe view_1" at 21,63 size 759x352
   TextField "Text field_1" at 309,10 size 209x27; Text 'Recipes Management / Recepie Management'
   GraphicView "Graphic view_61" at 2,4 size 149x43; Picture "logo2"
   DateTimeField "Date/time field_1" at 629,14 size 166x19
   Button "Button_1" at 6,432 size 88x38; TextOff 'Root'
      on Release: ActivateScreen("Root screen", 0)
      on Press: ActivateScreen("Root screen", 0)
   Button "Button_2" at 99,432 size 93x38; TextOff 'User / Benutzer'
      on Release: ActivateScreen("User administration", 0)
      on Press: ActivateScreen("User administration", 0)
   Button "Button_3" at 197,431 size 96x39; TextOff 'Alarms / Alarme'
      on Release: ActivateScreen("Alarm screen", 0)
      on Press: ActivateScreen("Alarm screen", 0)
   Button "Button_4" at 298,431 size 121x39; TextOff 'PLC diagnose / SPS Diagnose'
      on Release: ActivateScreen("SIMATIC PLC system diagnostics", 0)
      on Press: ActivateScreen("SIMATIC PLC system diagnostics", 0)
   Button "Button_5" at 425,431 size 106x39; TextOff 'Recipes / Rezepte'
      on Release: ActivateScreen("Recipes management", 0)
      on Press: ActivateScreen("Recipes management", 0)
   Button "Button_6" at 537,431 size 113x39; TextOff 'Visulization / Visulisierung'
      on Release: ActivateScreen("visualization", 0)
      on Press: ActivateScreen("visualization", 0)
   Button "Button_7" at 654,431 size 139x39; TextOff 'Historic Data / Frühere Daten'
      on Release: ActivateScreen("Historical Data", 0)
      on Press: ActivateScreen("Historical Data", 0)

screen "Engineer Screen" 800x480
   TextField "Text field_1" at 339,10 size 221x27; Text 'Engineer Screen / Gruppe der Ingenieure'
   GraphicView "Graphic view_61" at 2,4 size 149x43; Picture "logo2"
   DateTimeField "Date/time field_1" at 629,14 size 166x19
   Button "Button_1" at 6,386 size 101x36; TextOff 'Logoff / Abmeldung'
      on Release: function_f23ef4c9()
      on Press: function_f23ef4c9(); ActivateScreen("Root screen", 0)
   RecipeView "Recipe view_1" at 8,56 size 630x323
   Group "Group_1" at 676,104 size 102x224
   Button "Button_2" at 6,432 size 88x38; TextOff 'Root'
      on Release: ActivateScreen("Root screen", 0)
      on Press: ActivateScreen("Root screen", 0)
   Button "Button_3" at 99,432 size 93x38; TextOff 'User / Benutzer'
      on Release: ActivateScreen("User administration", 0)
      on Press: ActivateScreen("User administration", 0)
   Button "Button_4" at 197,431 size 96x39; TextOff 'Alarms / Alarme'
      on Release: ActivateScreen("Alarm screen", 0)
      on Press: ActivateScreen("Alarm screen", 0)
   Button "Button_5" at 298,431 size 121x39; TextOff 'PLC diagnose / SPS Diagnose'
      on Release: ActivateScreen("SIMATIC PLC system diagnostics", 0)
      on Press: ActivateScreen("SIMATIC PLC system diagnostics", 0)
   Button "Button_6" at 425,431 size 106x39; TextOff 'Recipes / Rezepte'
      on Release: ActivateScreen("Recipes management", 0)
      on Press: ActivateScreen("Recipes management", 0)
   Button "Button_7" at 537,431 size 113x39; TextOff 'Visulization / Visulisierung'
      on Release: ActivateScreen("visualization", 0)
      on Press: ActivateScreen("visualization", 0)
   Button "Button_8" at 654,431 size 139x39; TextOff 'Historic Data / Frühere Daten'
      on Release: ActivateScreen("Historical Data", 0)
      on Press: ActivateScreen("Historical Data", 0)
   IOField "I/O field_2" at 677,215 size 96x32; FormatPattern 99; Unit %
      ProcessValue <- "Global_DB_Other_Parameters_Liquid_B_pct"
   Group "Group" at 676,266 size 102x62
   TextField "Text field_3" at 684,183 size 89x23; Text 'Liquid B%'
   IOField "I/O field_1" at 677,134 size 96x32; FormatPattern 99; Unit %
      ProcessValue <- "Global_DB_Other_Parameters_Liquid_A_pct"
   TextField "Text field_2" at 678,104 size 90x23; Text 'Liquid A%'
   IOField "I/O field_3" at 676,296 size 102x32; FormatPattern 999.99; Unit ml/s
      ProcessValue <- "Flow_ml_per_sec"
   TextField "Text field_4" at 680,266 size 87x23; Text 'Flow Rate'

screen "Alarm screen" 800x480
   TextField "Text field_1" at 343,10 size 72x27; Text 'Alarms / Alarme'
   GraphicView "Graphic view_61" at 2,4 size 149x43; Picture "logo2"
   DateTimeField "Date/time field_1" at 629,14 size 166x19
   AlarmView "Alarm view_1" at 25,66 size 744x347
   Button "Button_1" at 6,432 size 88x38; TextOff 'Root'
      on Release: ActivateScreen("Root screen", 0)
      on Press: ActivateScreen("Root screen", 0)
   Button "Button_2" at 99,432 size 93x38; TextOff 'User / Benutzer'
      on Release: ActivateScreen("User administration", 0)
      on Press: ActivateScreen("User administration", 0)
   Button "Button_3" at 197,431 size 96x39; TextOff 'Alarms / Alarme'
      on Release: ActivateScreen("Alarm screen", 0)
      on Press: ActivateScreen("Alarm screen", 0)
   Button "Button_4" at 298,431 size 121x39; TextOff 'PLC diagnose / SPS Diagnose'
      on Release: ActivateScreen("SIMATIC PLC system diagnostics", 0)
      on Press: ActivateScreen("SIMATIC PLC system diagnostics", 0)
   Button "Button_5" at 425,431 size 106x39; TextOff 'Recipes / Rezepte'
      on Release: ActivateScreen("Recipes management", 0)
      on Press: ActivateScreen("Recipes management", 0)
   Button "Button_6" at 537,431 size 113x39; TextOff 'Visulization / Visulisierung'
      on Release: ActivateScreen("visualization", 0)
      on Press: ActivateScreen("visualization", 0)
   Button "Button_7" at 654,431 size 139x39; TextOff 'Historic Data / Frühere Daten'
      on Release: ActivateScreen("Historical Data", 0)
      on Press: ActivateScreen("Historical Data", 0)

Template "Template_1" 800x480
   Button "Template_Button" at 714,429 size 71x50; TextOff 'Text'
   Button "Template_Button_1" at 614,429 size 71x50; TextOff 'Text'
   Button "Template_Button_2" at 514,429 size 71x50; TextOff 'Text'
   Button "Template_Button_3" at 414,429 size 71x50; TextOff 'Text'
   Button "Template_Button_4" at 314,429 size 71x50; TextOff 'Text'
   Button "Template_Button_5" at 214,429 size 71x50; TextOff 'Text'
   Button "Template_Button_6" at 114,429 size 71x50; TextOff 'Text'
   Button "Alarms" at 14,429 size 71x50; TextOn 'Alarms / Alarme'; TextOff 'Alarms / Alarme'; PictureOn "AlarmDisplay_KTP700_Basic_DP_TR"; PictureOff "AlarmDisplay_KTP700_Basic_DP_TR"
      on Release: function_ef3f5d25("Alarm window_Unacknowledged", -1)
   DateTimeField "HmiScreenItemData" at 695,25 size 105x25
   DateTimeField "HmiScreenItemData_1" at 695,0 size 105x25
*)